      Contact( "14_DQ_DATA".CV_421_5S )
   END_RUNG wire#w1
   RUNG wire#w2
      Contact( "FIT417_5S_ALM_ANALOG_DB"."ALARM H" )
      Coil( %DB2062.DBX7.1 )
   END_RUNG
   // the same network as SCL:
   "FIT417_5S_ALM_ANALOG_DB"(Value := "20_TANKS_IP_DATA".RIO_05.SECOND_TANK.USD_FLOW,   // "502_ALM_ANALOG"
                           "Raw Value" := "Tank 5S USD Flow Meter",
                           Enable := "2100_AUTO_SEQ_DB".SEQ_RNG AND "14_DQ_DATA".CV_421_5S,
                           "SHORT CIRCUIT VALUE" := 32000.0,
                           "BROKEN WIRE VALUE" := -32000.0,
                           "VERY LOW LEVEL VALUE (LL)" := "2084_Setpoints".FIT418_LoLo,
                           "LOW LEVEL VALUE (L)" := "2084_Setpoints".FIT418_Lo,
                           "HIGH LEVEL VALUE (H)" := "2084_Setpoints".FIT418_Hi,
                           "VERY HIGH LEVEL VALUE (HH)" := "2084_Setpoints".FIT418_HiHi,
                           "ALARM DELAY" := "2086_Times"."FIT417STAR Alarm Delay",
                           "ALARM READING" => %DB2062.DBX363.4,
                           ENO => #_w1);
   %DB2062.DBX7.0 := #_w1 AND "FIT417_5S_ALM_ANALOG_DB"."ALARM L";
   %DB2062.DBX7.1 := #_w1 AND "FIT417_5S_ALM_ANALOG_DB"."ALARM H";
END_REGION

REGION Network 31: DB2062.DBX7.2 = FIT418 6Port USD Flow LO / DB2062.DBX7.3 = FIT418 6Port USD Flow HI
   // BTCS_WARNING_WORD_04_BIT_10/11                      12.13
   RUNG wire#powerrail
      "FIT418_6P__ALM_ANALOG_DB"(Enable := wire#w1, Value := "20_TANKS_IP_DATA".RIO_06.FIRST_TANK.USD_FLOW, "Raw Value" := "Tank 6P USD Flow Meter", "Enable Delay Time" :=, "High Value Release" :=, "SHORT CIRCUIT VALUE" := 32000.0, "BROKEN WIRE VALUE" := -32000.0, "VERY LOW LEVEL VALUE (LL)" := "2084_Setpoints".FIT418_LoLo, "LOW LEVEL VALUE (L)" := "2084_Setpoints".FIT418_Lo, "HIGH LEVEL VALUE (H)" := "2084_Setpoints".FIT418_Hi, "VERY HIGH LEVEL VALUE (HH)" := "2084_Setpoints".FIT418_HiHi, OFFSET :=, "ALARM DELAY" := "2086_Times"."FIT418PORT Alarm Delay", "Peak Value Reset" :=, "ALARM HH" =>, "ALARM H" =>, "ALARM L" =>, "ALARM LL" =>, "ALARM READING" => %DB2062.DBX363.5, "Peak Value" =>, Alarm =>, Alarm_INT =>)
      wire#w2
      Contact( "FIT418_6P__ALM_ANALOG_DB"."ALARM L" )
      Coil( %DB2062.DBX7.2 )
   END_RUNG
   RUNG wire#powerrail
      Contact( "2100_AUTO_SEQ_DB".SEQ_RNG )
      Contact( "14_DQ_DATA".CV_422_6P )
   END_RUNG wire#w1
   RUNG wire#w2
      Contact( "FIT418_6P__ALM_ANALOG_DB"."ALARM H" )
      Coil( %DB2062.DBX7.3 )
   END_RUNG
   // the same network as SCL:
   "FIT418_6P__ALM_ANALOG_DB"(Value := "20_TANKS_IP_DATA".RIO_06.FIRST_TANK.USD_FLOW,   // "502_ALM_ANALOG"
                           "Raw Value" := "Tank 6P USD Flow Meter",
                           Enable := "2100_AUTO_SEQ_DB".SEQ_RNG AND "14_DQ_DATA".CV_422_6P,
                           "SHORT CIRCUIT VALUE" := 32000.0,
                           "BROKEN WIRE VALUE" := -32000.0,
                           "VERY LOW LEVEL VALUE (LL)" := "2084_Setpoints".FIT418_LoLo,
                           "LOW LEVEL VALUE (L)" := "2084_Setpoints".FIT418_Lo,
                           "HIGH LEVEL VALUE (H)" := "2084_Setpoints".FIT418_Hi,
                           "VERY HIGH LEVEL VALUE (HH)" := "2084_Setpoints".FIT418_HiHi,
                           "ALARM DELAY" := "2086_Times"."FIT418PORT Alarm Delay",
                           "ALARM READING" => %DB2062.DBX363.5,
                           ENO => #_w1);
   %DB2062.DBX7.2 := #_w1 AND "FIT418_6P__ALM_ANALOG_DB"."ALARM L";
   %DB2062.DBX7.3 := #_w1 AND "FIT418_6P__ALM_ANALOG_DB"."ALARM H";
END_REGION

REGION Network 32: DB2062.DBX7.4 = FIT417 6Starboard USD Flow LO / DB2062.DBX7.5 = FIT417 6Starboard USD Flow HI
   // BTCS_WARNING_WORD_04_BIT_12/13                        12.14
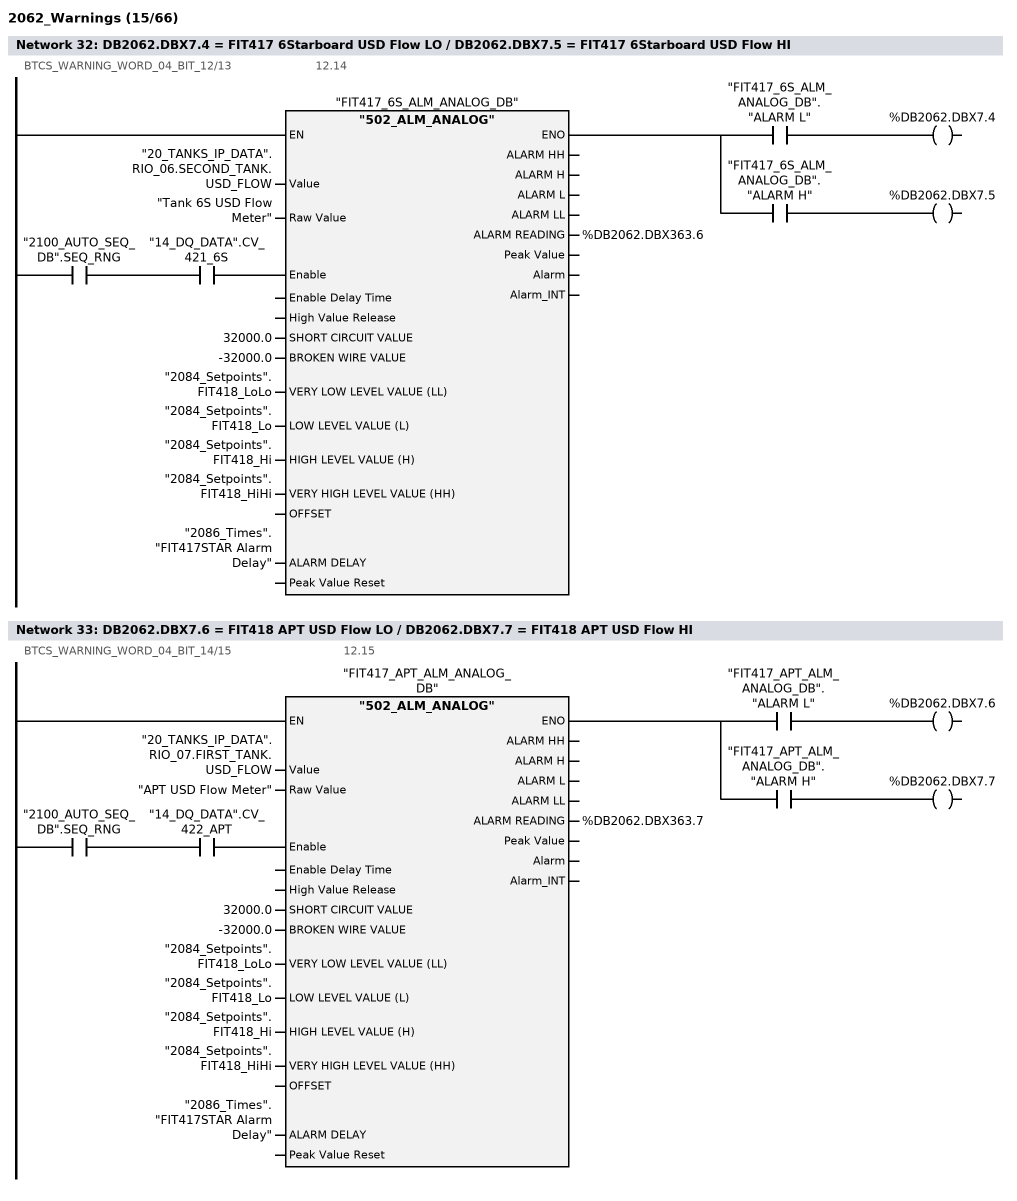
   RUNG wire#powerrail
      "FIT417_6S_ALM_ANALOG_DB"(Enable := wire#w1, Value := "20_TANKS_IP_DATA".RIO_06.SECOND_TANK.USD_FLOW, "Raw Value" := "Tank 6S USD Flow Meter", "Enable Delay Time" :=, "High Value Release" :=, "SHORT CIRCUIT VALUE" := 32000.0, "BROKEN WIRE VALUE" := -32000.0, "VERY LOW LEVEL VALUE (LL)" := "2084_Setpoints".FIT418_LoLo, "LOW LEVEL VALUE (L)" := "2084_Setpoints".FIT418_Lo, "HIGH LEVEL VALUE (H)" := "2084_Setpoints".FIT418_Hi, "VERY HIGH LEVEL VALUE (HH)" := "2084_Setpoints".FIT418_HiHi, OFFSET :=, "ALARM DELAY" := "2086_Times"."FIT417STAR Alarm Delay", "Peak Value Reset" :=, "ALARM HH" =>, "ALARM H" =>, "ALARM L" =>, "ALARM LL" =>, "ALARM READING" => %DB2062.DBX363.6, "Peak Value" =>, Alarm =>, Alarm_INT =>)
      wire#w2
      Contact( "FIT417_6S_ALM_ANALOG_DB"."ALARM L" )
      Coil( %DB2062.DBX7.4 )
   END_RUNG
   RUNG wire#powerrail
      Contact( "2100_AUTO_SEQ_DB".SEQ_RNG )
      Contact( "14_DQ_DATA".CV_421_6S )
   END_RUNG wire#w1
   RUNG wire#w2
      Contact( "FIT417_6S_ALM_ANALOG_DB"."ALARM H" )
      Coil( %DB2062.DBX7.5 )
   END_RUNG
   // the same network as SCL:
   "FIT417_6S_ALM_ANALOG_DB"(Value := "20_TANKS_IP_DATA".RIO_06.SECOND_TANK.USD_FLOW,   // "502_ALM_ANALOG"
                           "Raw Value" := "Tank 6S USD Flow Meter",
                           Enable := "2100_AUTO_SEQ_DB".SEQ_RNG AND "14_DQ_DATA".CV_421_6S,
                           "SHORT CIRCUIT VALUE" := 32000.0,
                           "BROKEN WIRE VALUE" := -32000.0,
                           "VERY LOW LEVEL VALUE (LL)" := "2084_Setpoints".FIT418_LoLo,
                           "LOW LEVEL VALUE (L)" := "2084_Setpoints".FIT418_Lo,
                           "HIGH LEVEL VALUE (H)" := "2084_Setpoints".FIT418_Hi,
                           "VERY HIGH LEVEL VALUE (HH)" := "2084_Setpoints".FIT418_HiHi,
                           "ALARM DELAY" := "2086_Times"."FIT417STAR Alarm Delay",
                           "ALARM READING" => %DB2062.DBX363.6,
                           ENO => #_w1);
   %DB2062.DBX7.4 := #_w1 AND "FIT417_6S_ALM_ANALOG_DB"."ALARM L";
   %DB2062.DBX7.5 := #_w1 AND "FIT417_6S_ALM_ANALOG_DB"."ALARM H";
END_REGION

REGION Network 33: DB2062.DBX7.6 = FIT418 APT USD Flow LO / DB2062.DBX7.7 = FIT418 APT USD Flow HI
   // BTCS_WARNING_WORD_04_BIT_14/15                                12.15
   RUNG wire#powerrail
      "FIT417_APT_ALM_ANALOG_DB"(Enable := wire#w1, Value := "20_TANKS_IP_DATA".RIO_07.FIRST_TANK.USD_FLOW, "Raw Value" := "APT USD Flow Meter", "Enable Delay Time" :=, "High Value Release" :=, "SHORT CIRCUIT VALUE" := 32000.0, "BROKEN WIRE VALUE" := -32000.0, "VERY LOW LEVEL VALUE (LL)" := "2084_Setpoints".FIT418_LoLo, "LOW LEVEL VALUE (L)" := "2084_Setpoints".FIT418_Lo, "HIGH LEVEL VALUE (H)" := "2084_Setpoints".FIT418_Hi, "VERY HIGH LEVEL VALUE (HH)" := "2084_Setpoints".FIT418_HiHi, OFFSET :=, "ALARM DELAY" := "2086_Times"."FIT417STAR Alarm Delay", "Peak Value Reset" :=, "ALARM HH" =>, "ALARM H" =>, "ALARM L" =>, "ALARM LL" =>, "ALARM READING" => %DB2062.DBX363.7, "Peak Value" =>, Alarm =>, Alarm_INT =>)
      wire#w2
      Contact( "FIT417_APT_ALM_ANALOG_DB"."ALARM L" )
      Coil( %DB2062.DBX7.6 )
   END_RUNG
   RUNG wire#powerrail
      Contact( "2100_AUTO_SEQ_DB".SEQ_RNG )
      Contact( "14_DQ_DATA".CV_422_APT )
   END_RUNG wire#w1
   RUNG wire#w2
      Contact( "FIT417_APT_ALM_ANALOG_DB"."ALARM H" )
      Coil( %DB2062.DBX7.7 )
   END_RUNG
   // the same network as SCL:
   "FIT417_APT_ALM_ANALOG_DB"(Value := "20_TANKS_IP_DATA".RIO_07.FIRST_TANK.USD_FLOW,   // "502_ALM_ANALOG"
                           "Raw Value" := "APT USD Flow Meter",
                           Enable := "2100_AUTO_SEQ_DB".SEQ_RNG AND "14_DQ_DATA".CV_422_APT,
                           "SHORT CIRCUIT VALUE" := 32000.0,
                           "BROKEN WIRE VALUE" := -32000.0,
                           "VERY LOW LEVEL VALUE (LL)" := "2084_Setpoints".FIT418_LoLo,
                           "LOW LEVEL VALUE (L)" := "2084_Setpoints".FIT418_Lo,
                           "HIGH LEVEL VALUE (H)" := "2084_Setpoints".FIT418_Hi,
                           "VERY HIGH LEVEL VALUE (HH)" := "2084_Setpoints".FIT418_HiHi,
                           "ALARM DELAY" := "2086_Times"."FIT417STAR Alarm Delay",
                           "ALARM READING" => %DB2062.DBX363.7,
                           ENO => #_w1);
   %DB2062.DBX7.6 := #_w1 AND "FIT417_APT_ALM_ANALOG_DB"."ALARM L";
   %DB2062.DBX7.7 := #_w1 AND "FIT417_APT_ALM_ANALOG_DB"."ALARM H";
END_REGION

REGION Network 35: DB2062.DBX8.0 = FIT420 FPT MBG Flow LO / DB2062.DBX8.1 = FIT420 FPT MBG Flow HI
   // BTCS_WARNING_WORD_05_BIT_0/1              13.0
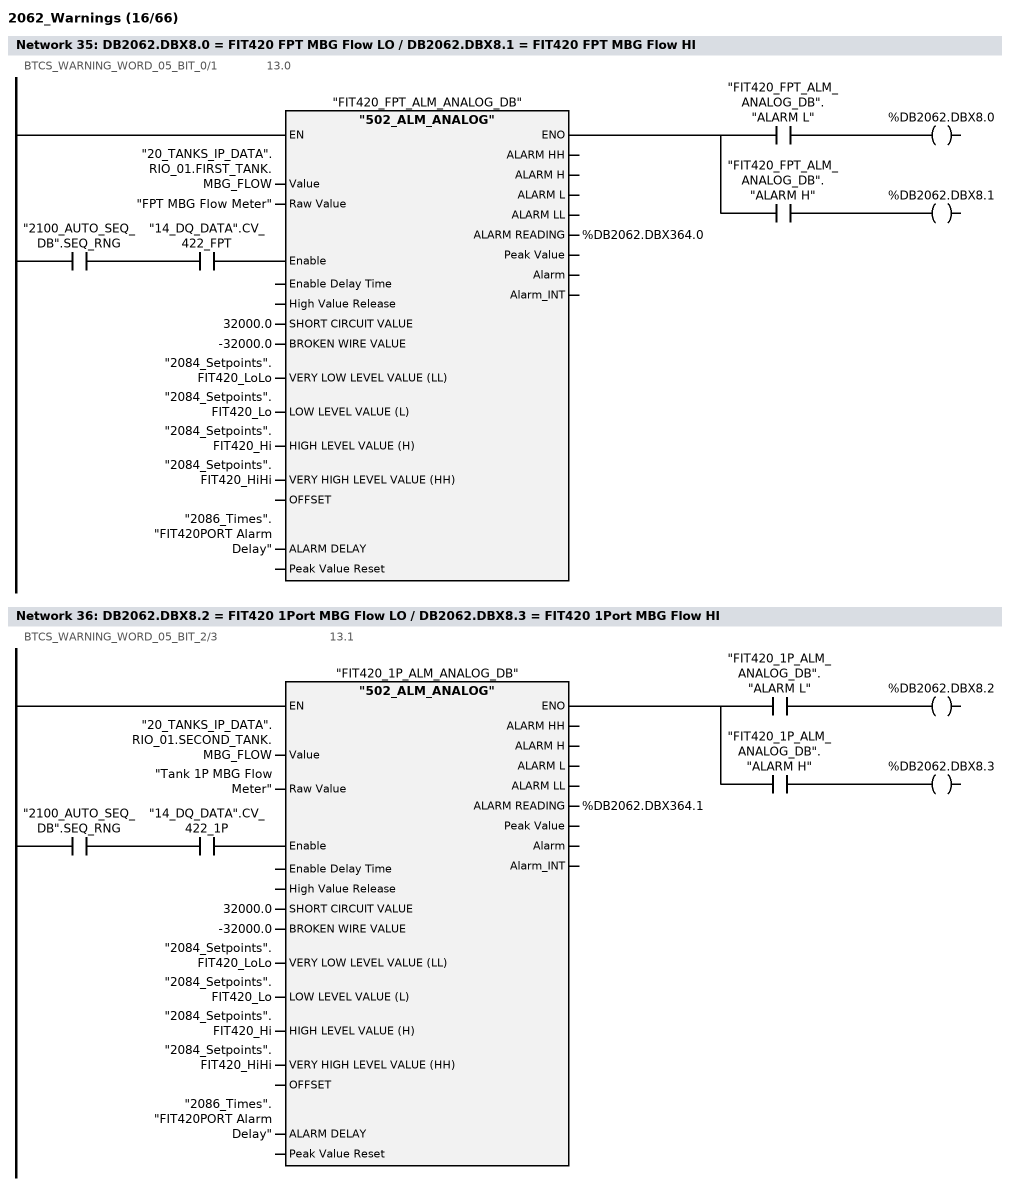
   RUNG wire#powerrail
      "FIT420_FPT_ALM_ANALOG_DB"(Enable := wire#w1, Value := "20_TANKS_IP_DATA".RIO_01.FIRST_TANK.MBG_FLOW, "Raw Value" := "FPT MBG Flow Meter", "Enable Delay Time" :=, "High Value Release" :=, "SHORT CIRCUIT VALUE" := 32000.0, "BROKEN WIRE VALUE" := -32000.0, "VERY LOW LEVEL VALUE (LL)" := "2084_Setpoints".FIT420_LoLo, "LOW LEVEL VALUE (L)" := "2084_Setpoints".FIT420_Lo, "HIGH LEVEL VALUE (H)" := "2084_Setpoints".FIT420_Hi, "VERY HIGH LEVEL VALUE (HH)" := "2084_Setpoints".FIT420_HiHi, OFFSET :=, "ALARM DELAY" := "2086_Times"."FIT420PORT Alarm Delay", "Peak Value Reset" :=, "ALARM HH" =>, "ALARM H" =>, "ALARM L" =>, "ALARM LL" =>, "ALARM READING" => %DB2062.DBX364.0, "Peak Value" =>, Alarm =>, Alarm_INT =>)
      wire#w2
      Contact( "FIT420_FPT_ALM_ANALOG_DB"."ALARM L" )
      Coil( %DB2062.DBX8.0 )
   END_RUNG
   RUNG wire#powerrail
      Contact( "2100_AUTO_SEQ_DB".SEQ_RNG )
      Contact( "14_DQ_DATA".CV_422_FPT )
   END_RUNG wire#w1
   RUNG wire#w2
      Contact( "FIT420_FPT_ALM_ANALOG_DB"."ALARM H" )
      Coil( %DB2062.DBX8.1 )
   END_RUNG
   // the same network as SCL:
   "FIT420_FPT_ALM_ANALOG_DB"(Value := "20_TANKS_IP_DATA".RIO_01.FIRST_TANK.MBG_FLOW,   // "502_ALM_ANALOG"
                           "Raw Value" := "FPT MBG Flow Meter",
                           Enable := "2100_AUTO_SEQ_DB".SEQ_RNG AND "14_DQ_DATA".CV_422_FPT,
                           "SHORT CIRCUIT VALUE" := 32000.0,
                           "BROKEN WIRE VALUE" := -32000.0,
                           "VERY LOW LEVEL VALUE (LL)" := "2084_Setpoints".FIT420_LoLo,
                           "LOW LEVEL VALUE (L)" := "2084_Setpoints".FIT420_Lo,
                           "HIGH LEVEL VALUE (H)" := "2084_Setpoints".FIT420_Hi,
                           "VERY HIGH LEVEL VALUE (HH)" := "2084_Setpoints".FIT420_HiHi,
                           "ALARM DELAY" := "2086_Times"."FIT420PORT Alarm Delay",
                           "ALARM READING" => %DB2062.DBX364.0,
                           ENO => #_w1);
   %DB2062.DBX8.0 := #_w1 AND "FIT420_FPT_ALM_ANALOG_DB"."ALARM L";
   %DB2062.DBX8.1 := #_w1 AND "FIT420_FPT_ALM_ANALOG_DB"."ALARM H";
END_REGION

REGION Network 36: DB2062.DBX8.2 = FIT420 1Port MBG Flow LO / DB2062.DBX8.3 = FIT420 1Port MBG Flow HI
   // BTCS_WARNING_WORD_05_BIT_2/3                                13.1
   RUNG wire#powerrail
      "FIT420_1P_ALM_ANALOG_DB"(Enable := wire#w1, Value := "20_TANKS_IP_DATA".RIO_01.SECOND_TANK.MBG_FLOW, "Raw Value" := "Tank 1P MBG Flow Meter", "Enable Delay Time" :=, "High Value Release" :=, "SHORT CIRCUIT VALUE" := 32000.0, "BROKEN WIRE VALUE" := -32000.0, "VERY LOW LEVEL VALUE (LL)" := "2084_Setpoints".FIT420_LoLo, "LOW LEVEL VALUE (L)" := "2084_Setpoints".FIT420_Lo, "HIGH LEVEL VALUE (H)" := "2084_Setpoints".FIT420_Hi, "VERY HIGH LEVEL VALUE (HH)" := "2084_Setpoints".FIT420_HiHi, OFFSET :=, "ALARM DELAY" := "2086_Times"."FIT420PORT Alarm Delay", "Peak Value Reset" :=, "ALARM HH" =>, "ALARM H" =>, "ALARM L" =>, "ALARM LL" =>, "ALARM READING" => %DB2062.DBX364.1, "Peak Value" =>, Alarm =>, Alarm_INT =>)
      wire#w2
      Contact( "FIT420_1P_ALM_ANALOG_DB"."ALARM L" )
      Coil( %DB2062.DBX8.2 )
   END_RUNG
   RUNG wire#powerrail
      Contact( "2100_AUTO_SEQ_DB".SEQ_RNG )
      Contact( "14_DQ_DATA".CV_422_1P )
   END_RUNG wire#w1
   RUNG wire#w2
      Contact( "FIT420_1P_ALM_ANALOG_DB"."ALARM H" )
      Coil( %DB2062.DBX8.3 )
   END_RUNG
   // the same network as SCL:
   "FIT420_1P_ALM_ANALOG_DB"(Value := "20_TANKS_IP_DATA".RIO_01.SECOND_TANK.MBG_FLOW,   // "502_ALM_ANALOG"
                           "Raw Value" := "Tank 1P MBG Flow Meter",
                           Enable := "2100_AUTO_SEQ_DB".SEQ_RNG AND "14_DQ_DATA".CV_422_1P,
                           "SHORT CIRCUIT VALUE" := 32000.0,
                           "BROKEN WIRE VALUE" := -32000.0,
                           "VERY LOW LEVEL VALUE (LL)" := "2084_Setpoints".FIT420_LoLo,
                           "LOW LEVEL VALUE (L)" := "2084_Setpoints".FIT420_Lo,
                           "HIGH LEVEL VALUE (H)" := "2084_Setpoints".FIT420_Hi,
                           "VERY HIGH LEVEL VALUE (HH)" := "2084_Setpoints".FIT420_HiHi,
                           "ALARM DELAY" := "2086_Times"."FIT420PORT Alarm Delay",
                           "ALARM READING" => %DB2062.DBX364.1,
                           ENO => #_w1);
   %DB2062.DBX8.2 := #_w1 AND "FIT420_1P_ALM_ANALOG_DB"."ALARM L";
   %DB2062.DBX8.3 := #_w1 AND "FIT420_1P_ALM_ANALOG_DB"."ALARM H";
END_REGION

REGION Network 37: DB2062.DBX8.4 = FIT419 1Starboard MBG Flow LO / DB2062.DBX8.5 = FIT419 1Starboard MBG Flow HI
   // BTCS_WARNING_WORD_05_BIT_4/5                      13.2
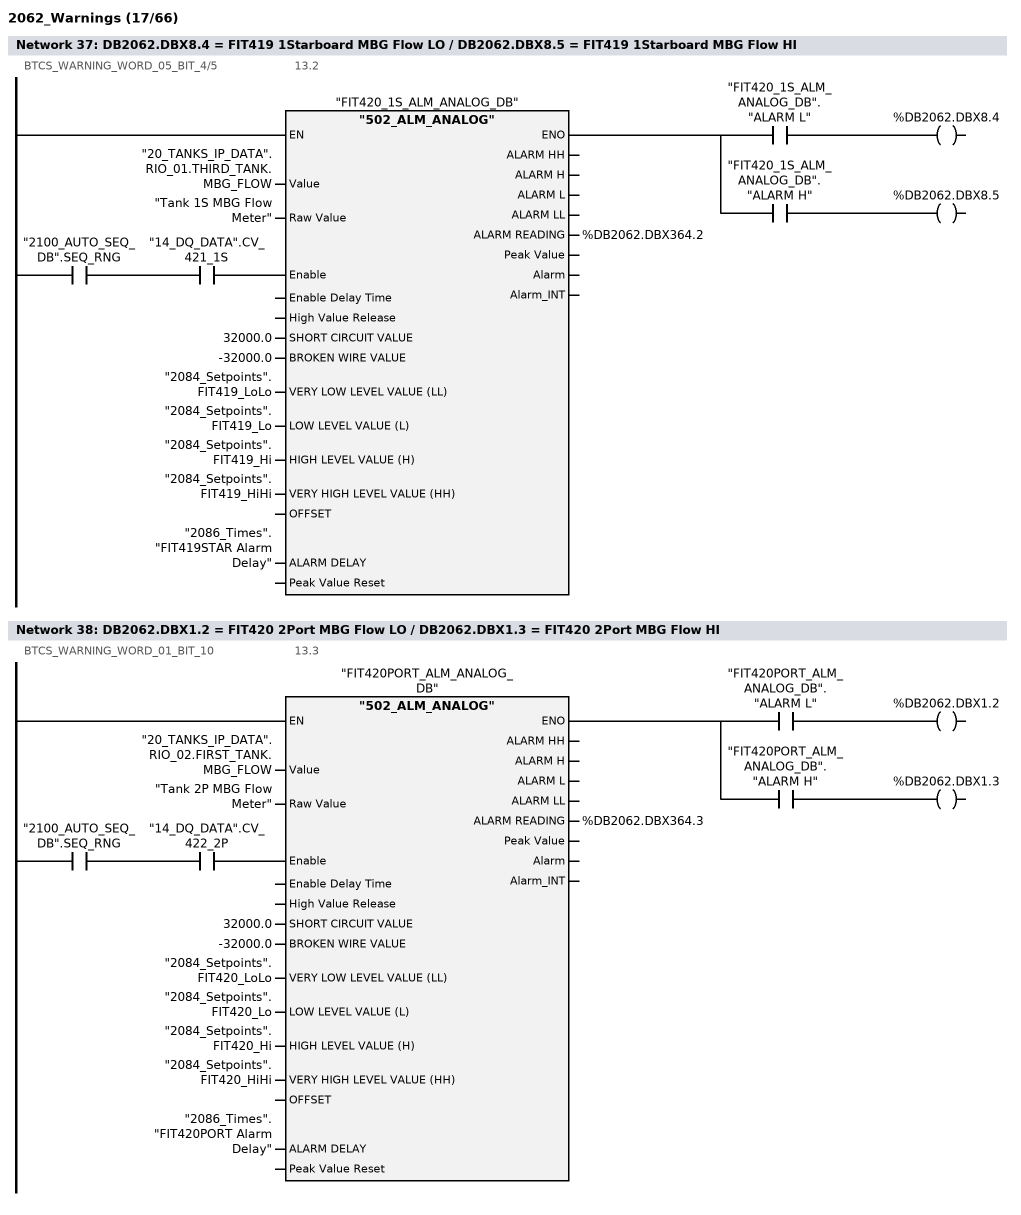
   RUNG wire#powerrail
      "FIT420_1S_ALM_ANALOG_DB"(Enable := wire#w1, Value := "20_TANKS_IP_DATA".RIO_01.THIRD_TANK.MBG_FLOW, "Raw Value" := "Tank 1S MBG Flow Meter", "Enable Delay Time" :=, "High Value Release" :=, "SHORT CIRCUIT VALUE" := 32000.0, "BROKEN WIRE VALUE" := -32000.0, "VERY LOW LEVEL VALUE (LL)" := "2084_Setpoints".FIT419_LoLo, "LOW LEVEL VALUE (L)" := "2084_Setpoints".FIT419_Lo, "HIGH LEVEL VALUE (H)" := "2084_Setpoints".FIT419_Hi, "VERY HIGH LEVEL VALUE (HH)" := "2084_Setpoints".FIT419_HiHi, OFFSET :=, "ALARM DELAY" := "2086_Times"."FIT419STAR Alarm Delay", "Peak Value Reset" :=, "ALARM HH" =>, "ALARM H" =>, "ALARM L" =>, "ALARM LL" =>, "ALARM READING" => %DB2062.DBX364.2, "Peak Value" =>, Alarm =>, Alarm_INT =>)
      wire#w2
      Contact( "FIT420_1S_ALM_ANALOG_DB"."ALARM L" )
      Coil( %DB2062.DBX8.4 )
   END_RUNG
   RUNG wire#powerrail
      Contact( "2100_AUTO_SEQ_DB".SEQ_RNG )
      Contact( "14_DQ_DATA".CV_421_1S )
   END_RUNG wire#w1
   RUNG wire#w2
      Contact( "FIT420_1S_ALM_ANALOG_DB"."ALARM H" )
      Coil( %DB2062.DBX8.5 )
   END_RUNG
   // the same network as SCL:
   "FIT420_1S_ALM_ANALOG_DB"(Value := "20_TANKS_IP_DATA".RIO_01.THIRD_TANK.MBG_FLOW,   // "502_ALM_ANALOG"
                           "Raw Value" := "Tank 1S MBG Flow Meter",
                           Enable := "2100_AUTO_SEQ_DB".SEQ_RNG AND "14_DQ_DATA".CV_421_1S,
                           "SHORT CIRCUIT VALUE" := 32000.0,
                           "BROKEN WIRE VALUE" := -32000.0,
                           "VERY LOW LEVEL VALUE (LL)" := "2084_Setpoints".FIT419_LoLo,
                           "LOW LEVEL VALUE (L)" := "2084_Setpoints".FIT419_Lo,
                           "HIGH LEVEL VALUE (H)" := "2084_Setpoints".FIT419_Hi,
                           "VERY HIGH LEVEL VALUE (HH)" := "2084_Setpoints".FIT419_HiHi,
                           "ALARM DELAY" := "2086_Times"."FIT419STAR Alarm Delay",
                           "ALARM READING" => %DB2062.DBX364.2,
                           ENO => #_w1);
   %DB2062.DBX8.4 := #_w1 AND "FIT420_1S_ALM_ANALOG_DB"."ALARM L";
   %DB2062.DBX8.5 := #_w1 AND "FIT420_1S_ALM_ANALOG_DB"."ALARM H";
END_REGION

REGION Network 38: DB2062.DBX1.2 = FIT420 2Port MBG Flow LO / DB2062.DBX1.3 = FIT420 2Port MBG Flow HI
   // BTCS_WARNING_WORD_01_BIT_10                       13.3
   RUNG wire#powerrail
      "FIT420PORT_ALM_ANALOG_DB"(Enable := wire#w1, Value := "20_TANKS_IP_DATA".RIO_02.FIRST_TANK.MBG_FLOW, "Raw Value" := "Tank 2P MBG Flow Meter", "Enable Delay Time" :=, "High Value Release" :=, "SHORT CIRCUIT VALUE" := 32000.0, "BROKEN WIRE VALUE" := -32000.0, "VERY LOW LEVEL VALUE (LL)" := "2084_Setpoints".FIT420_LoLo, "LOW LEVEL VALUE (L)" := "2084_Setpoints".FIT420_Lo, "HIGH LEVEL VALUE (H)" := "2084_Setpoints".FIT420_Hi, "VERY HIGH LEVEL VALUE (HH)" := "2084_Setpoints".FIT420_HiHi, OFFSET :=, "ALARM DELAY" := "2086_Times"."FIT420PORT Alarm Delay", "Peak Value Reset" :=, "ALARM HH" =>, "ALARM H" =>, "ALARM L" =>, "ALARM LL" =>, "ALARM READING" => %DB2062.DBX364.3, "Peak Value" =>, Alarm =>, Alarm_INT =>)
      wire#w2
      Contact( "FIT420PORT_ALM_ANALOG_DB"."ALARM L" )
      Coil( %DB2062.DBX1.2 )
   END_RUNG
   RUNG wire#powerrail
      Contact( "2100_AUTO_SEQ_DB".SEQ_RNG )
      Contact( "14_DQ_DATA".CV_422_2P )
   END_RUNG wire#w1
   RUNG wire#w2
      Contact( "FIT420PORT_ALM_ANALOG_DB"."ALARM H" )
      Coil( %DB2062.DBX1.3 )
   END_RUNG
   // the same network as SCL:
   "FIT420PORT_ALM_ANALOG_DB"(Value := "20_TANKS_IP_DATA".RIO_02.FIRST_TANK.MBG_FLOW,   // "502_ALM_ANALOG"
                           "Raw Value" := "Tank 2P MBG Flow Meter",
                           Enable := "2100_AUTO_SEQ_DB".SEQ_RNG AND "14_DQ_DATA".CV_422_2P,
                           "SHORT CIRCUIT VALUE" := 32000.0,
                           "BROKEN WIRE VALUE" := -32000.0,
                           "VERY LOW LEVEL VALUE (LL)" := "2084_Setpoints".FIT420_LoLo,
                           "LOW LEVEL VALUE (L)" := "2084_Setpoints".FIT420_Lo,
                           "HIGH LEVEL VALUE (H)" := "2084_Setpoints".FIT420_Hi,
                           "VERY HIGH LEVEL VALUE (HH)" := "2084_Setpoints".FIT420_HiHi,
                           "ALARM DELAY" := "2086_Times"."FIT420PORT Alarm Delay",
                           "ALARM READING" => %DB2062.DBX364.3,
                           ENO => #_w1);
   %DB2062.DBX1.2 := #_w1 AND "FIT420PORT_ALM_ANALOG_DB"."ALARM L";
   %DB2062.DBX1.3 := #_w1 AND "FIT420PORT_ALM_ANALOG_DB"."ALARM H";
END_REGION

REGION Network 39: DB2062.DBX1.6 = FIT419 2Starboard MBG Flow LO / DB2062.DBX1.7 = FIT419 2Starboard MBG Flow HI
   // BTCS_WARNING_WORD_01_BIT_14                          13.4
